(* CODESYS project Revisora_V2.0.1f.project (continued)
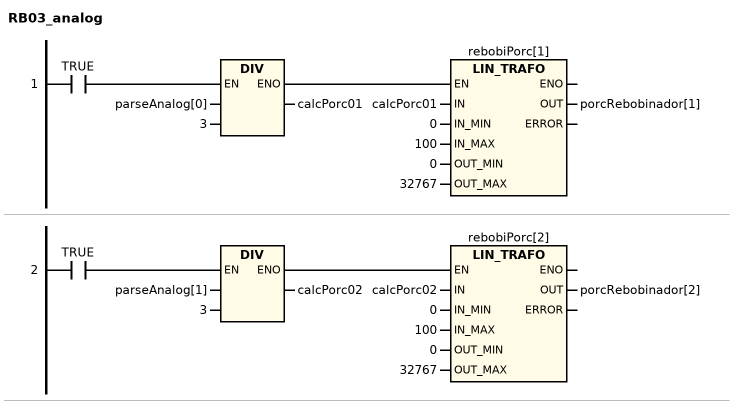
// NETWORK 1
calcPorc01 := parseAnalog[0] / 3;
rebobiPorc[1](
    IN := calcPorc01,
    IN_MIN := 0,
    IN_MAX := 100,
    OUT_MIN := 0,
    OUT_MAX := 32767,
    OUT => porcRebobinador[1]); // LIN_TRAFO

// NETWORK 2
calcPorc02 := parseAnalog[1] / 3;
rebobiPorc[2](
    IN := calcPorc02,
    IN_MIN := 0,
    IN_MAX := 100,
    OUT_MIN := 0,
    OUT_MAX := 32767,
    OUT => porcRebobinador[2]); // LIN_TRAFO

END_PROGRAM

// MyController/Application/02_Rebobinadores/RB04_saidas
PROGRAM RB04_saidas
VAR
END_VAR

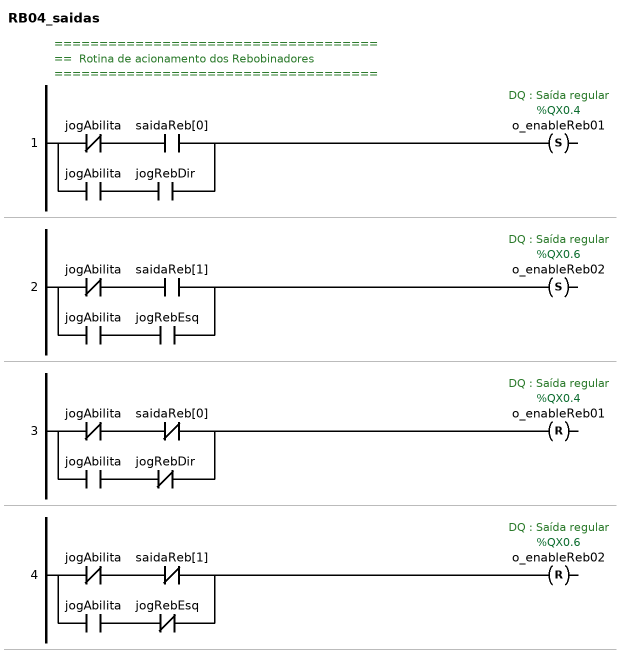
// NETWORK 1
// ====================================
// ==  Rotina de acionamento dos Rebobinadores
// ====================================
//   o_enableReb01: DQ : Saída regular | AT %QX0.4
o_enableReb01 S= NOT jogAbilita AND saidaReb[0] OR jogAbilita AND jogRebDir;

// NETWORK 2
//   o_enableReb02: DQ : Saída regular | AT %QX0.6
o_enableReb02 S= NOT jogAbilita AND saidaReb[1] OR jogAbilita AND jogRebEsq;

// NETWORK 3
//   o_enableReb01: DQ : Saída regular | AT %QX0.4
o_enableReb01 R= NOT jogAbilita AND NOT saidaReb[0] OR jogAbilita AND NOT jogRebDir;

// NETWORK 4
//   o_enableReb02: DQ : Saída regular | AT %QX0.6
o_enableReb02 R= NOT jogAbilita AND NOT saidaReb[1] OR jogAbilita AND NOT jogRebEsq;

END_PROGRAM

// MyController/Application/02_Rebobinadores/RB05_sentido
PROGRAM RB05_sentido
VAR
auxParseAnalog				:ARRAY [1..2] OF REAL;
END_VAR

// Calcula quando o valor for menor que 0
auxParseAnalog[1]:= (parseAnalog[0] * 328) / 3;
auxParseAnalog[2]:= (parseAnalog[1] * 328) / 3;

IF parseAnalog[0] < 0 THEN
	valorPorcRebobinador[1]:= auxParseAnalog[1];
ELSE
	valorPorcRebobinador[1]:= porcRebobinador[1];	
END_IF

IF parseAnalog[1] < 0 THEN
	valorPorcRebobinador[2]:= auxParseAnalog[2];
ELSE
	valorPorcRebobinador[2]:= porcRebobinador[2];	
END_IF

// Sentido dos rebobinadores
IF	enbReb.IP THEN
	IF i_sentido THEN
		ladoDir:= FALSE;
		ladoEsq:= TRUE;
		visLadoEsq:= TRUE;
		visLadoDir:= FALSE;
		displayState:= 0;
	ELSE
		ladoEsq:= FALSE;
		ladoDir:= TRUE;
		visLadoEsq:= FALSE;
		visLadoDir:= TRUE;
		displayState:= 1;
	END_IF
END_IF

// Editar valores

	IF ladoEsq THEN
		analoReb02:= REAL_TO_INT((valorPorcRebobinador[1])*-1); 
		analoReb01:= REAL_TO_INT((valorPorcRebobinador[2]));
		delayTorq[0] := T#0MS;
		delayTorq[1] := T#90MS;
		
	END_IF
	
	IF ladoDir THEN
		analoReb02:= REAL_TO_INT(valorPorcRebobinador[2])*-1;
		analoReb01:= REAL_TO_INT(valorPorcRebobinador[1]);
		delayTorq[0] := T#90MS;
		delayTorq[1] := T#0MS;
	END_IF
	
	//IF NOT ciclo.IP THEN
	//	ladoEsq:= FALSE;
	//	ladoDir:= FALSE;
//	END_IF
	
	// Parada
	IF torqueParada THEN
		IF ladoEsq THEN
			analoReb01:= -1311;
			analoReb02:= -1311;
		ELSE
			analoReb01:= 1311;
			analoReb02:= 1311;
		END_IF
	END_IF
// Calcula quando o valor for menor que 0
//auxParseAnalog[1]:= (parseAnalog[0] * 328) / 3;
//auxParseAnalog[2]:= (parseAnalog[1] * 328) / 3;

END_PROGRAM

// MyController/Application/03_Nip/NP01_geral
PROGRAM NP01_geral
VAR
	TD_power				: TOF;
END_VAR
VAR // added by the converter: edge detectors and wires of the graphical bodies
    _ft1 : F_TRIG;
END_VAR

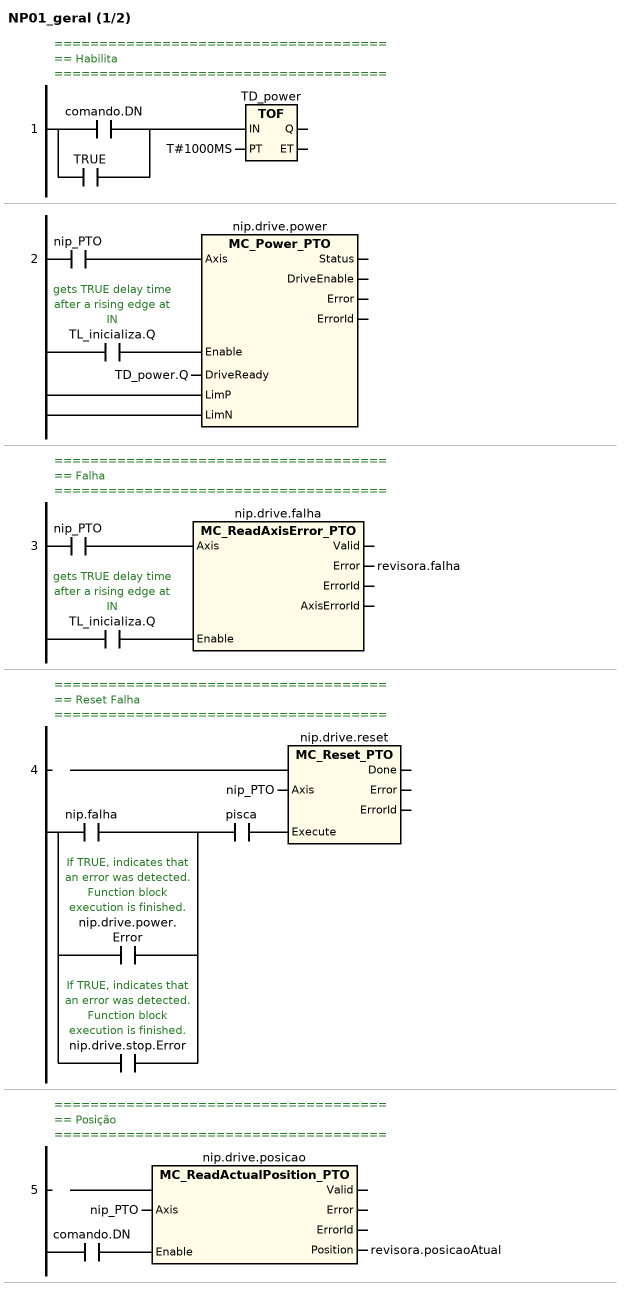
// NETWORK 1
// =====================================
// == Habilita
// =====================================
TD_power(IN := comando.DN OR TRUE, PT := T#1000MS); // TOF

// NETWORK 2
//   TL_inicializa.Q: gets TRUE delay time after a rising edge at IN
//   TD_power.Q: gets FALSE, when PT milliseconds elapsed, since falling edge at IN
nip.drive.power(
    Axis := nip_PTO,
    Enable := TL_inicializa.Q,
    DriveReady := TD_power.Q,
    LimP := TRUE,
    LimN := TRUE); // MC_Power_PTO

// NETWORK 3
// =====================================
// == Falha
// =====================================
//   TL_inicializa.Q: gets TRUE delay time after a rising edge at IN
nip.drive.falha(Axis := nip_PTO, Enable := TL_inicializa.Q, Error => revisora.falha); // MC_ReadAxisError_PTO

// NETWORK 4
// =====================================
// == Reset Falha
// =====================================
//   nip.drive.power.Error: If TRUE, indicates that an error was detected. Function block execution is finished.
//   nip.drive.stop.Error: If TRUE, indicates that an error was detected. Function block execution is finished.
nip.drive.reset(Axis := nip_PTO, Execute := (nip.falha OR nip.drive.power.Error OR nip.drive.stop.Error) AND pisca); // MC_Reset_PTO

// NETWORK 5
// =====================================
// == Posição
// =====================================
nip.drive.posicao(Axis := nip_PTO, Enable := comando.DN, Position => revisora.posicaoAtual); // MC_ReadActualPosition_PTO

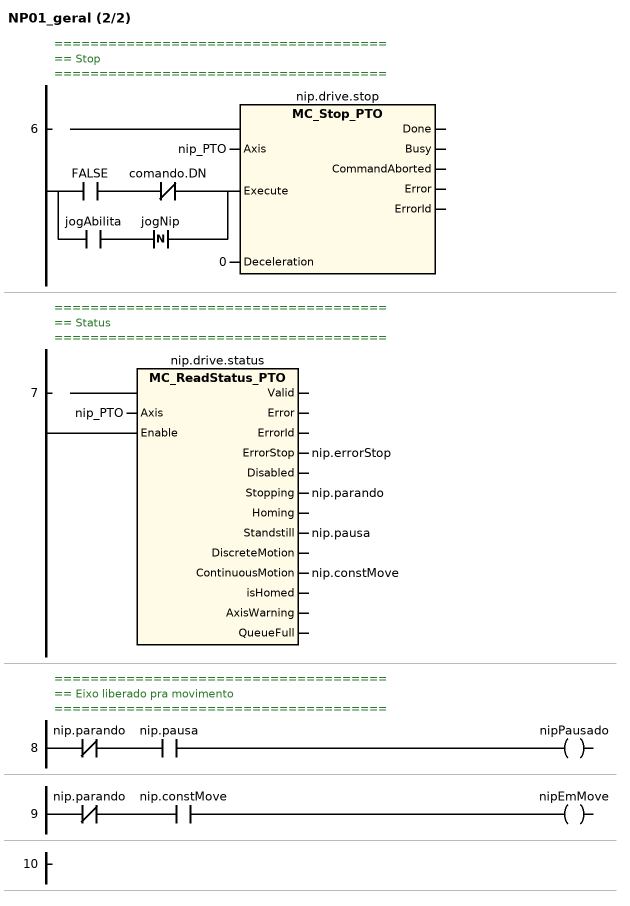
// NETWORK 6
// =====================================
// == Stop
// =====================================
_ft1(CLK := jogNip);
nip.drive.stop(
    Axis := nip_PTO,
    Execute := FALSE AND NOT comando.DN OR jogAbilita AND _ft1.Q,
    Deceleration := 0); // MC_Stop_PTO

// NETWORK 7
// =====================================
// == Status
// =====================================
nip.drive.status(
    Axis := nip_PTO,
    Enable := TRUE,
    ErrorStop => nip.errorStop,
    Stopping => nip.parando,
    Standstill => nip.pausa,
    ContinuousMotion => nip.constMove); // MC_ReadStatus_PTO

// NETWORK 8
// =====================================
// == Eixo liberado pra movimento
// =====================================
nipPausado := NOT nip.parando AND nip.pausa;

// NETWORK 9
nipEmMove := NOT nip.parando AND nip.constMove;

// NETWORK 10

END_PROGRAM

// MyController/Application/03_Nip/NP02_enableNip
PROGRAM NP02_enableNip
VAR
END_VAR

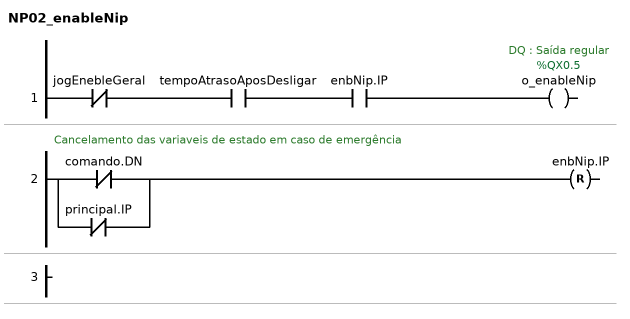
// NETWORK 1
//   o_enableNip: DQ : Saída regular | AT %QX0.5
o_enableNip := NOT jogEnebleGeral AND tempoAtrasoAposDesligar AND enbNip.IP;

// NETWORK 2
// Cancelamento das variaveis de estado em caso de emergência
enbNip.IP R= NOT comando.DN OR NOT principal.IP;

// NETWORK 3

END_PROGRAM

// MyController/Application/03_Nip/NP03_auto
PROGRAM NP03_auto
VAR
	TF_enable						: TON;
	MC_MoveVelocity_PTO_0			: MC_MoveVelocity_PTO;
	atrasoAposDesligar				: TON;
END_VAR
VAR // added by the converter: edge detectors and wires of the graphical bodies
    _rt1 : R_TRIG;
    _ft1, _ft2 : F_TRIG;
    _w1, _w2 : BOOL;
END_VAR

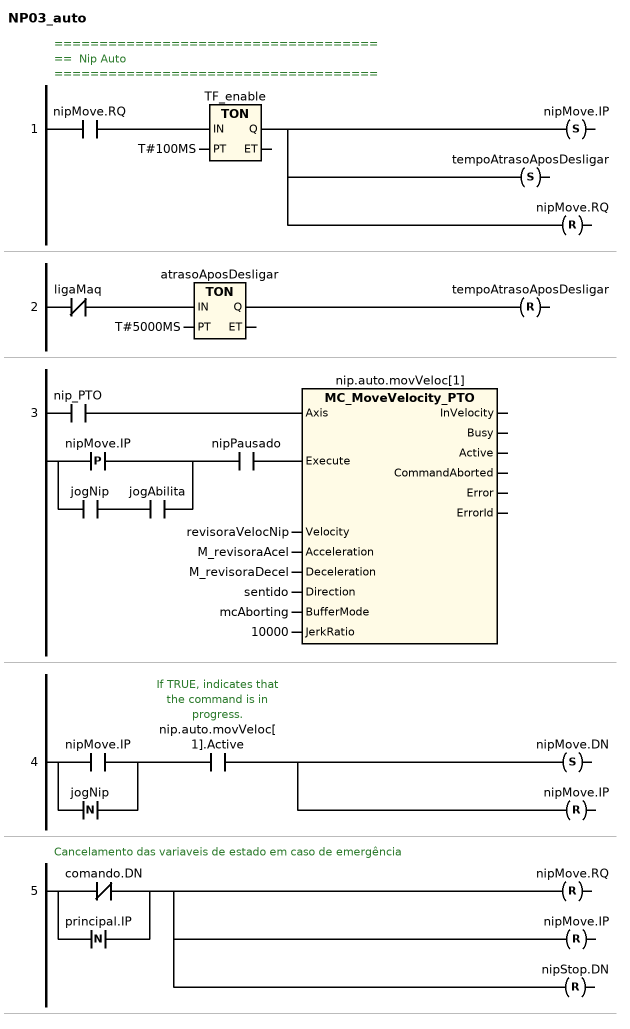
// NETWORK 1
// ====================================
// ==  Nip Auto
// ====================================
TF_enable(IN := nipMove.RQ, PT := T#100MS); // TON
nipMove.IP S= TF_enable.Q;
tempoAtrasoAposDesligar S= TF_enable.Q;
nipMove.RQ R= TF_enable.Q;

// NETWORK 2
atrasoAposDesligar(IN := NOT ligaMaq, PT := T#5000MS); // TON
tempoAtrasoAposDesligar R= atrasoAposDesligar.Q;

// NETWORK 3
_rt1(CLK := nipMove.IP);
nip.auto.movVeloc[1](
    Axis := nip_PTO,
    Execute := (_rt1.Q OR jogNip AND jogAbilita) AND nipPausado,
    Velocity := revisoraVelocNip,
    Acceleration := M_revisoraAcel,
    Deceleration := M_revisoraDecel,
    Direction := sentido,
    BufferMode := mcAborting,
    JerkRatio := 10000); // MC_MoveVelocity_PTO

// NETWORK 4
//   nip.auto.movVeloc[1].Active: If TRUE, indicates that the command is in progress.
_ft1(CLK := jogNip);
_w1 := (nipMove.IP OR _ft1.Q) AND nip.auto.movVeloc[1].Active;
nipMove.DN S= _w1;
nipMove.IP R= _w1;

// NETWORK 5
// Cancelamento das variaveis de estado em caso de emergência
_ft2(CLK := principal.IP);
_w2 := NOT comando.DN OR _ft2.Q;
nipMove.RQ R= _w2;
nipMove.IP R= _w2;
nipStop.DN R= _w2;

END_PROGRAM

// MyController/Application/03_Nip/NP04_parada
PROGRAM NP04_parada
VAR
	testeFW			: BOOL;
	job: BOOL;
END_VAR
VAR // added by the converter: edge detectors and wires of the graphical bodies
    _w1, _w2, _w3 : BOOL;
    _rt1 : R_TRIG;
    _ft1 : F_TRIG;
END_VAR

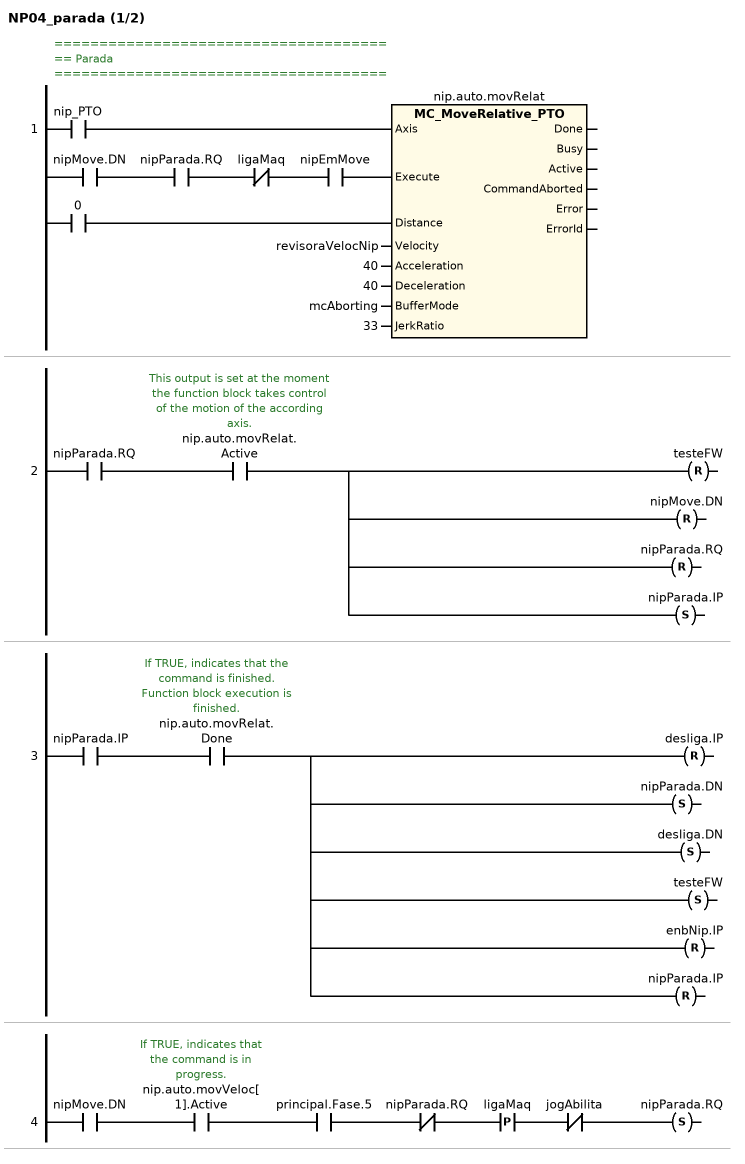
// NETWORK 1
// =====================================
// == Parada
// =====================================
nip.auto.movRelat(
    Axis := nip_PTO,
    Execute := nipMove.DN AND nipParada.RQ AND NOT ligaMaq AND nipEmMove,
    Distance := 0,
    Velocity := revisoraVelocNip,
    Acceleration := 40,
    Deceleration := 40,
    BufferMode := mcAborting,
    JerkRatio := 33); // MC_MoveRelative_PTO

// NETWORK 2
//   nip.auto.movRelat.Active: This output is set at the moment the function block takes control of the motion of the according axis.
_w1 := nipParada.RQ AND nip.auto.movRelat.Active;
testeFW R= _w1;
nipMove.DN R= _w1;
nipParada.RQ R= _w1;
nipParada.IP S= _w1;

// NETWORK 3
//   nip.auto.movRelat.Done: If TRUE, indicates that the command is finished. Function block execution is finished.
_w2 := nipParada.IP AND nip.auto.movRelat.Done;
desliga.IP R= _w2;
nipParada.DN S= _w2;
desliga.DN S= _w2;
testeFW S= _w2;
enbNip.IP R= _w2;
nipParada.IP R= _w2;

// NETWORK 4
//   nip.auto.movVeloc[1].Active: If TRUE, indicates that the command is in progress.
_rt1(CLK := ligaMaq);
nipParada.RQ S= nipMove.DN AND nip.auto.movVeloc[1].Active AND principal.Fase.5 AND NOT nipParada.RQ AND _rt1.Q AND NOT jogAbilita;

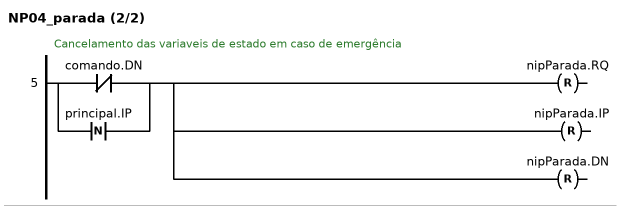
// NETWORK 5
// Cancelamento das variaveis de estado em caso de emergência
_ft1(CLK := principal.IP);
_w3 := NOT comando.DN OR _ft1.Q;
nipParada.RQ R= _w3;
nipParada.IP R= _w3;
nipParada.DN R= _w3;

END_PROGRAM

// MyController/Application/03_Nip/NP06_jog
PROGRAM NP06_jog
VAR
	auxJogPos								: BOOL;
	auxJopNeg								: BOOL;
END_VAR
VAR // added by the converter: edge detectors and wires of the graphical bodies
    _ft1, _ft2 : F_TRIG;
END_VAR

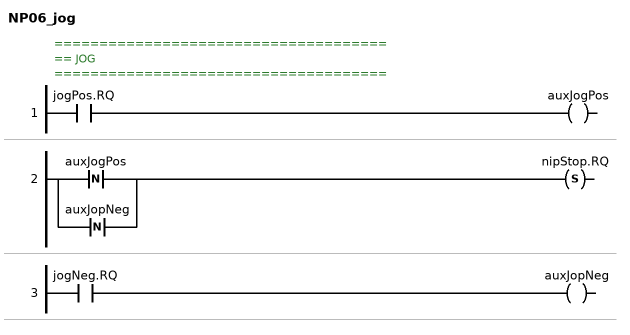
// NETWORK 1
// =====================================
// == JOG
// =====================================
auxJogPos := jogPos.RQ;

// NETWORK 2
_ft1(CLK := auxJogPos);
_ft2(CLK := auxJopNeg);
nipStop.RQ S= _ft1.Q OR _ft2.Q;

// NETWORK 3
auxJopNeg := jogNeg.RQ;

END_PROGRAM

// MyController/Application/03_Nip/NP07_veloc
PROGRAM NP07_veloc
VAR

	timerVeloc 		: TON;

END_VAR

// Partida Lenta
M_revisoraVeloc:=bobinaAtual.velocReb;
//IF nipMove.RQ THEN
//	IF bobinaAtual.velocDesb > 800 OR bobinaAtual.velocReb > 800 THEN	
	//	M_revisoraVeloc:= 600;
	//	partidaLenta:= TRUE;
//	END_IF
//END_IF

//timerVeloc(IN:= partidaLenta, PT:= T#7S);

//IF 	timerVeloc.Q THEN
	//nipMove.IP:= FALSE;
	//partidaLenta:= FALSE;
	//IF i_sentido THEN
	//	M_revisoraVeloc:= bobinaAtual.velocDesb;
	//	nipMove.IP:= TRUE;
//	ELSE
//		M_revisoraVeloc:= bobinaAtual.velocReb;
//		nipMove.IP:= TRUE;
//	END_IF
//END_IF

//IF NOT comando.DN OR principal.IP OR ligaMaq THEN
//	partidaLenta:= FALSE;
//END_IF

END_PROGRAM

// MyController/Application/03_Nip/NP09_sentido
PROGRAM NP09_sentido
VAR
END_VAR

// Mudança de sentido
IF i_sentido AND NOT ciclo.IP THEN
	sentido:= 1;
	M_pulsosParar:= 20;
ELSIF NOT i_sentido AND NOT ciclo.IP THEN
	sentido:= -1;
	M_pulsosParar:= -20;
END_IF

END_PROGRAM

// MyController/Application/03_Nip/NP20_JogTest
PROGRAM NP20_JogTest
VAR
	auxVeloc			:DINT;
	auxReb01			: INT;
	auxReb02			: INT;
END_VAR

IF jogVelocNip >3000 THEN
	jogVelocNip:= 3000;
	
END_IF

IF jogAbilita = TRUE THEN
	revisoraVelocNip:=jogVelocNip;
ELSE
	revisoraVelocNip:=M_revisoraVeloc;
END_IF

END_PROGRAM

// MyController/Application/05_IHM/I01_geral
PROGRAM I01_geral
VAR
	auxBit				: BOOL;
END_VAR
VAR // added by the converter: edge detectors and wires of the graphical bodies
    _rt1 : R_TRIG;
END_VAR

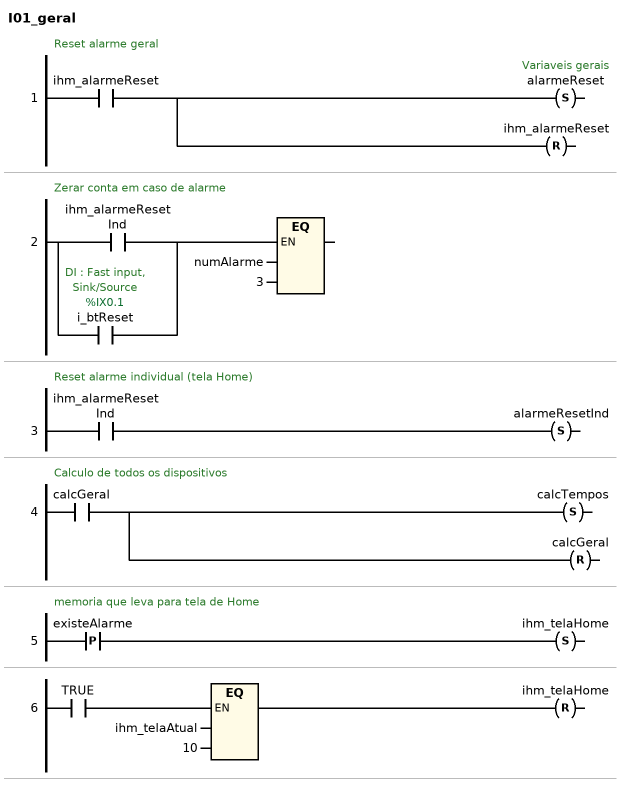
// NETWORK 1
// Reset alarme geral
//   alarmeReset: Variaveis gerais
alarmeReset S= ihm_alarmeReset;
ihm_alarmeReset R= ihm_alarmeReset;

// NETWORK 2
// Zerar conta em caso de alarme
//   i_btReset: DI : Fast input, Sink/Source | AT %IX0.1
(* (ihm_alarmeResetInd OR i_btReset) AND numAlarme = 3; result not used *)

// NETWORK 3
// Reset alarme individual (tela Home)
alarmeResetInd S= ihm_alarmeResetInd;

// NETWORK 4
// Calculo de todos os dispositivos
calcTempos S= calcGeral;
calcGeral R= calcGeral;

// NETWORK 5
// memoria que leva para tela de Home
_rt1(CLK := existeAlarme);
ihm_telaHome S= _rt1.Q;

// NETWORK 6
ihm_telaHome R= ihm_telaAtual = 10;

END_PROGRAM

// MyController/Application/05_IHM/I02_alarmes
PROGRAM I02_alarmes
VAR
	auxExisteAlarme					: BOOL;
	delayAlarme						: TON;
	memAlarme						: ARRAY[0..99] OF BOOL;
	p0								: SINT;
END_VAR


CASE alarmes.Fase OF
(*====================================
  ==  Fase 0 - alarmes 1 a 50 (0 não existe)
  ====================================*)
0:
	auxExisteAlarme:= FALSE;
	FOR p0:= 1 TO 50 DO
		IF alarme[p0] THEN
			memAlarme[p0]:= TRUE;
			auxExisteAlarme:= TRUE;
			
			IF numAlarme = 0 THEN
				numAlarme:= p0;				// pega o numero do primeiro alarme que ocorre
			END_IF
		END_IF
		
		IF numAlarme = p0 THEN
			IF alarme[p0] = 0 THEN			// verifica se o alarme que ocorreu continua ativo
				numAlarme:= 0;
			END_IF
		END_IF
	END_FOR
	alarmes.Fase:= 10;

	
(*====================================
  ==  Fase 10 - passa alarmes para ihm	
  ====================================*)
10:
	FOR p0:= 1 TO 50 DO
		ihm_alarme[p0]:= memAlarme[p0];
		memAlarme[p0]:= FALSE;
	END_FOR
	alarmes.Fase:= 11;
	
	
(*====================================
  ==  Fase 11 - verifica cancela alarmes pela IHM
  ====================================*)	
11:
	existeAlarme:= auxExisteAlarme;
	IF alarmeReset THEN
		alarmes.Fase:= 12;
	ELSE
		IF alarmeResetInd OR (i_btReset AND comando.DN) THEN
			alarme[numAlarme]:= FALSE;
			alarmeResetInd:= FALSE;
		END_IF
		alarmes.Fase:= 0;
	END_IF

	
(*====================================
  ==  Fase 12 - cancela alarmes	
  ====================================*)
12:
	alarmeReset:= FALSE;
	FOR p0:= 1 TO 50 DO
		alarme[p0]:= 0;
	END_FOR
	alarmes.Fase:= 13;
	

(*====================================
  ==  Fase 13 - espera 100ms para atualização dos bits de alarmes pelo controle
  ====================================*)	
13:
	IF delayAlarme.Q THEN
		alarmes.Fase:= 0;
	END_IF
	delayAlarme(IN:= alarmes.Fase= 13, PT:= T#100MS);

END_CASE

END_PROGRAM

// MyController/Application/05_IHM/I03_mensagens
PROGRAM I03_mensagens
VAR
	delayMensag						: TON;
	mensagens						: _exec_bits;
	p1								: DINT;
END_VAR


IF NOT mensagens.RQ THEN
	FOR p1:= 1 TO 50 DO
		IF mensagem[p1] = TRUE THEN
			mensagem[p1]:= 0;
			ihm_mensagem:= p1;
			mensagens.RQ:= TRUE;
		END_IF
	END_FOR
END_IF


// Tempo de cada mensagem na tela
delayMensag(IN := ihm_bannerMensagem, PT:= T#2500MS);
IF delayMensag.Q THEN
	mensagens.RQ:= FALSE;
	ihm_mensagem:= 0;
END_IF


ihm_bannerMensagem:= mensagens.RQ AND NOT ihm_bannerConfirma;

END_PROGRAM

// MyController/Application/05_IHM/I06_textoConfirma
PROGRAM I06_textoConfirma
VAR
END_VAR
VAR // added by the converter: edge detectors and wires of the graphical bodies
    _w1 : BOOL;
END_VAR

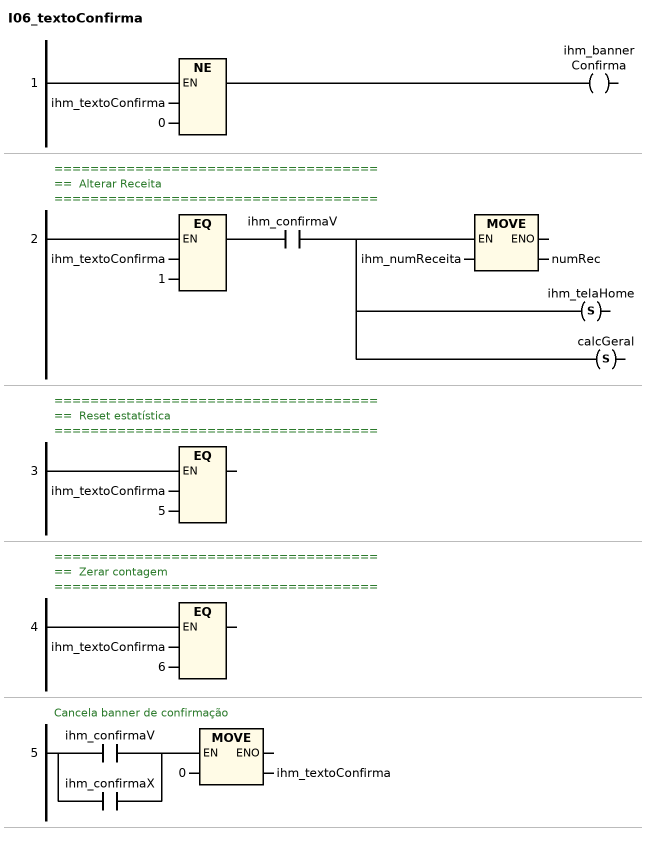
// NETWORK 1
ihm_bannerConfirma := ihm_textoConfirma <> 0;

// NETWORK 2
// ====================================
// ==  Alterar Receita
// ====================================
_w1 := ihm_textoConfirma = 1 AND ihm_confirmaV;
IF _w1 THEN numRec := ihm_numReceita; END_IF
ihm_telaHome S= _w1;
calcGeral S= _w1;

// NETWORK 3
// ====================================
// ==  Reset estatística
// ====================================
(* ihm_textoConfirma = 5; result not used *)

// NETWORK 4
// ====================================
// ==  Zerar contagem
// ====================================
(* ihm_textoConfirma = 6; result not used *)

// NETWORK 5
// Cancela banner de confirmação
IF ihm_confirmaV OR ihm_confirmaX THEN ihm_textoConfirma := 0; END_IF

END_PROGRAM

// MyController/Application/10_Relogio/AjustaDataHora
PROGRAM AjustaDataHora
VAR
	writeDateTime			: SetDateAndTime;
	readDateTime			: GetDateAndTime;
	bitScan					: BOOL;
	comOk					: BOOL;
	T_com					: TON;
END_VAR
VAR // added by the converter: edge detectors and wires of the graphical bodies
    _rt1 : R_TRIG;
END_VAR

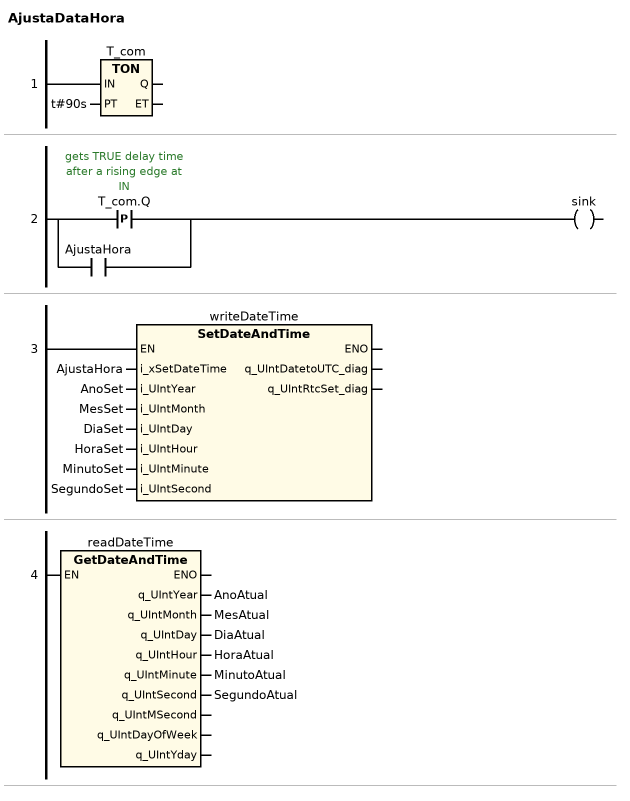
// NETWORK 1
T_com(IN := TRUE, PT := t#90s); // TON

// NETWORK 2
//   T_com.Q: gets TRUE delay time after a rising edge at IN
_rt1(CLK := T_com.Q);
sink := _rt1.Q OR AjustaHora;

// NETWORK 3
//   AnoSet: Sincroniza e ajusta o relógio da IHM
writeDateTime(
    i_xSetDateTime := AjustaHora,
    i_UIntYear := AnoSet,
    i_UIntMonth := MesSet,
    i_UIntDay := DiaSet,
    i_UIntHour := HoraSet,
    i_UIntMinute := MinutoSet,
    i_UIntSecond := SegundoSet); // SetDateAndTime

// NETWORK 4
readDateTime(
    q_UIntYear => AnoAtual,
    q_UIntMonth => MesAtual,
    q_UIntDay => DiaAtual,
    q_UIntHour => HoraAtual,
    q_UIntMinute => MinutoAtual,
    q_UIntSecond => SegundoAtual); // GetDateAndTime

END_PROGRAM

// MyController/Application/10_Relogio/SetDateAndTime
FUNCTION_BLOCK SetDateAndTime
VAR_INPUT
	i_xSetDateTime			: BOOL; (* seta novo horário na transição false para true*)
	i_UIntYear				: UINT:=2011; (*Valor para o ano a ser ajustado*)
	i_UIntMonth				: UINT:=1;(*Valor para o mes a ser ajustado*) 
	i_UIntDay				: UINT:=1;(*Valor para o dia a ser ajustado*) 
	i_UIntHour				: UINT:=0; (*Valor para a hora a ser ajustada*)
	i_UIntMinute			: UINT:=0; (*Valor para o minuto a ser ajustado*)
	i_UIntSecond			: UINT:=0;(*Valor para o segundo a ser ajustado*)
END_VAR
VAR_OUTPUT
	q_UIntDatetoUTC_diag	: UDINT; (*Status quando se =0 ok se <>0 erro nas informações de entrada*)
	q_UIntRtcSet_diag		: UDINT; (*Status quando se =0 ok se <>0 erro nas informações de entrada*)
END_VAR
VAR
	My_UTC					: DWORD; 
	MyDateTime				: SYSTIMEDATE; 
	milesec					: UINT:=0;
	dayOfWeek				: UINT:=1;
	yday					: UINT:=1;
END_VAR
VAR // added by the converter: edge detectors and wires of the graphical bodies
    _s1 : SYSTIMEDATE;
    _w1, _w2 : ANY;
END_VAR

// compose _s1 : SYSTIMEDATE
_s1.wYear := i_UIntYear;
_s1.wMonth := i_UIntMonth;
_s1.wDay := i_UIntDay;
_s1.wHour := i_UIntHour;
_s1.wMinute := i_UIntMinute;
_s1.wSecond := i_UIntSecond;
_s1.wMilliseconds := milesec;
_s1.wDayOfWeek := dayOfWeek;
_s1.wYday := yday;
MyDateTime := _s1;
_w1 := SysTimeRtcConvertDateToUtc(pDate := MyDateTime, pdwTimestampUtc := My_UTC);
q_UIntDatetoUTC_diag := _w1;
IF My_UTC <> 16#FFFFFFFF AND i_xSetDateTime THEN _w2 := SysTimeRtcSet(ulTimestamp := My_UTC); END_IF
q_UIntRtcSet_diag := _w2;
i_xSetDateTime := FALSE;

END_FUNCTION_BLOCK

// MyController/Application/10_Relogio/GetDateAndTime
FUNCTION_BLOCK GetDateAndTime
VAR_INPUT
END_VAR
VAR_OUTPUT
	q_UIntYear			: UINT; 
	q_UIntMonth			: UINT; 
	q_UIntDay			: UINT; 
	q_UIntHour			: UINT; 
	q_UIntMinute		: UINT; 
	q_UIntSecond		: UINT; 
	q_UIntMSecond		: UINT; 
	q_UIntDayOfWeek		: UINT; 
	q_UIntYday			: UINT;
END_VAR
VAR
	Ctrl_DateTime		: SYSTIMEDATE; 
	// SysTimeRtcGet operation diag 
	GetTimeResult		: UDINT; 
// SysTimeRtcConvertUtcToDate operation diag 
	UTCtoDate_diag		: UDINT; 
END_VAR
VAR // added by the converter: edge detectors and wires of the graphical bodies
    _w1, _w2 : ANY;
END_VAR

_w1 := SysTimeRtcGet(pResult := GetTimeResult);
_w2 := SysTimeRtcConvertUtcToDate(dwTimestampUtc := _w1, pDate := Ctrl_DateTime);
UTCtoDate_diag := _w2;
q_UIntYear := Ctrl_DateTime.SYSTIMEDATE;
q_UIntMonth := Ctrl_DateTime.wYear;
q_UIntDay := Ctrl_DateTime.wMonth;
q_UIntHour := Ctrl_DateTime.wDay;
q_UIntMinute := Ctrl_DateTime.wHour;
q_UIntSecond := Ctrl_DateTime.wMinute;
q_UIntMSecond := Ctrl_DateTime.wSecond;
q_UIntDayOfWeek := Ctrl_DateTime.wMilliseconds;
q_UIntYday := Ctrl_DateTime.wDayOfWeek;

END_FUNCTION_BLOCK

// MyController/Application/02_Rebobinadores/RB01_enableReb
PROGRAM RB01_enableReb
VAR
	TL_Rebobinadores 			 	: TON;
	TL_delayTorque					: ARRAY [0..1] OF TON;
	auxDesligaReb					: BOOL;
END_VAR
VAR // added by the converter: edge detectors and wires of the graphical bodies
    _rt1 : R_TRIG;
    _ft1 : F_TRIG;
    _w1 : BOOL;
END_VAR

